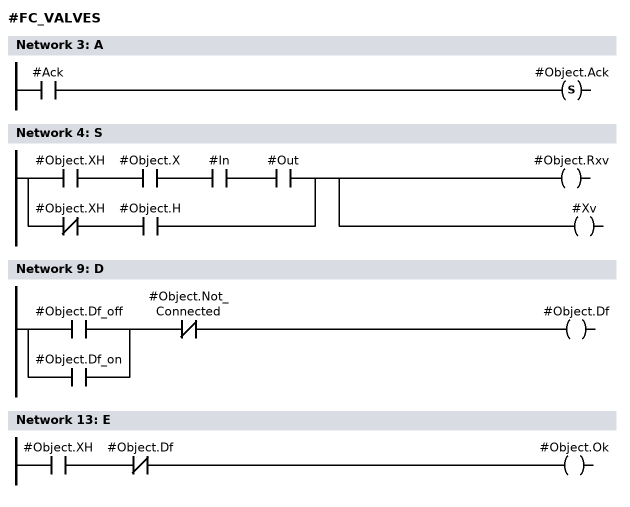
   RUNG wire#powerrail
      Contact( #Ack )
      S_Coil( #Object.Ack )
   END_RUNG
   // the same network as SCL:
   IF #Ack THEN #Object.Ack := TRUE; END_IF;
END_REGION

REGION Network 4: S
   RUNG wire#powerrail
      Contact( #Object.XH )
      Contact( #Object.X )
      Contact( #In )
      Contact( #Out )
      wire#w1
      Coil( #Object.Rxv )
   END_RUNG
   RUNG wire#powerrail
      I_Contact( #Object.XH )
      Contact( #Object.H )
   END_RUNG wire#w1
   RUNG wire#w1
      Coil( #Xv )
   END_RUNG
   // the same network as SCL:
   #Object.Rxv := (#Object.XH AND #Object.X AND #In AND #Out) OR (NOT #Object.XH AND #Object.H);
   #Xv := #Object.Rxv;
END_REGION

REGION Network 5 (STL): M
         A     #Object.XH;
         A     #Object.Rxv;
         S     #Object.H;

         A     #Object.XH;
         AN    #Object.Rxv;
         R     #Object.H;
END_REGION

REGION Network 6 (STL): R
         O(;
         AN    #Object.Inh;
         A     #Zs_on;
         );
         O(;
         A     #Object.Inh;
         A     #Object.Rxv;
         );
         =     #Object.Rzson;


         O(;
         AN    #Object.Inh;
         A     #Zs_off;
         );
         O(;
         A     #Object.Inh;
         AN    #Object.Rxv;
         );
         =     #Object.Rzsoff;


         AN    #In;
         =     #Object.R_in;


         AN    #Out;
         =     #Object.R_out;
END_REGION

REGION Network 7 (STL): D
         A     #Object.Rxv;
         A(;
         A(;
         ON    #Object.Rzson;
         O(;
         A     #Object.Rzsoff;
         A     #Object.Rzson;
         );
         );
         O(;
         A     #Object.Df_on;
         AN    #Object.Ack;
         );
         );
         =     #Temp1;


         CALL  "#FC_TIMER"
         ( Input     := #Temp1,
           Input_RTZ := FALSE,
           Pulse     := "point1secPls",
           RTZ       := FALSE,
           Tbase     := 1,
           Preset1   := #dTime,
           Preset2   := #Object.Gen.Para.Preset_Df_on,
           Time1     := #dTime,
           Time2     := #Object.Internal.Df_on
         );



         AN    #Object.Df_on;
         A(;
         L     #Object.Internal.Df_on;
         L     #Object.Gen.Para.Preset_Df_on;
         ==D;
         );
         JC    FON5;
         JU    FON6;
   FON5: S     #Object.Df_on;


   FON6: A     #Object.Ack;
         JC    FON7;
         JU    FON8;
   FON7: L     0;
         T     #Object.Internal.Df_on;
         R     #Object.Df_on;
   FON8: NOP   0;
END_REGION

REGION Network 8 (STL): d
         AN    #Object.Rxv;
         A(;
         O(;
         ON    #Object.Rzsoff;
         O(;
         A     #Object.Rzsoff;
         A     #Object.Rzson;
         );
         );
         O(;
         A     #Object.Df_off;
         AN    #Object.Ack;
         );
         );
         =     #Temp2;



         CALL  "#FC_TIMER"
         ( Input     := #Temp2,
           Input_RTZ := FALSE,
           Pulse     := "point1secPls",
           RTZ       := FALSE,
           Tbase     := 1,
           Preset1   := #dTime,
           Preset2   := #Object.Gen.Para.Preset_Df_off,
           Time1     := #dTime,
           Time2     := #Object.Internal.Df_off
         );


         AN    #Object.Df_off;
         A(;
         L     #Object.Internal.Df_off;
         L     #Object.Gen.Para.Preset_Df_off;
         ==D;
         );
         JC    FOF5;
         JU    FOF6;
   FOF5: S     #Object.Df_off;


   FOF6: A     #Object.Ack;
         JC    FOF7;
         JU    FOF8;
   FOF7: L     0;
         T     #Object.Internal.Df_off;
         R     #Object.Df_off;
   FOF8: NOP   0;
END_REGION

REGION Network 9: D
   RUNG wire#powerrail
      Contact( #Object.Df_off )
      wire#w1
      I_Contact( #Object.Not_Connected )
      Coil( #Object.Df )
   END_RUNG
   RUNG wire#powerrail
      Contact( #Object.Df_on )
   END_RUNG wire#w1
   // the same network as SCL:
   #Object.Df := (#Object.Df_off OR #Object.Df_on) AND NOT #Object.Not_Connected;
END_REGION

REGION Network 10 (STL): C
         A     #Object.Rxv;
         =     #Object.Internal.X_re_counter;

         CALL  "#FC_COUNTER"
         ( Input    := #Object.Internal.X_re_counter,
           Fr_input := #Object.Internal.Re_counter,
           Raz      := #Object.Raz_Fct_Run,
           Count    := #Object.C_run
         );
END_REGION

REGION Network 11 (STL): T
         CALL  "#FC_TIMER"
         ( Input     := #Object.Internal.X_re_counter,
           Input_RTZ := #Object.Raz_Fct_Run,
           Pulse     := "oneSecPls",
           RTZ       := TRUE,
           Tbase     := 1,
           Preset1   := 2073600000,
           Preset2   := #tTime,
           Time1     := #Object.T_run,
           Time2     := #tTime
         );
END_REGION

REGION Network 12 (STL): I
         CALL  "#FC_INH"
         ( Para_inh   := #Object.Gen.Para.Preset_T_exp_inh,
           Object_inh := #Object.Inh,
           Fe_inh     := #Object.Internal.Fe_inh,
           T_inh      := #Object.Internal.T_exp_inh
         );
END_REGION

REGION Network 13: E
   RUNG wire#powerrail
      Contact( #Object.XH )
      I_Contact( #Object.Df )
      Coil( #Object.Ok )
   END_RUNG
   // the same network as SCL:
   #Object.Ok := #Object.XH AND NOT #Object.Df;
END_REGION

REGION Network 14 (STL): Epics State
   // Copy of Auto/Manual mode
         A     #Object.XH;
         =     #sEpics.sAuto;

   // Copy of Inhibition mode
         A     #Object.Inh;
         =     #sEpics.sSim;

   // Copy of Command
         A     #Object.Rxv;
         =     #sEpics.sCmd;

   // Copy of On sensor
         A     #Object.Rzson;
         =     #sEpics.sOn;

   // Copy of Off sensor
         A     #Object.Rzsoff;
         =     #sEpics.sOff;

   // Copy of On fault
         A     #Object.Df_on;
         =     #sEpics.sOnFlt;

   // Copy of Off fault
         A     #Object.Df_off;
         =     #sEpics.sOffFlt;

   // Copy of Faults
         O     #Object.Df_on;
         O     #Object.Df_off;
         =     #sEpics.sFlt;

   // Copy of Command in Auto
         A     #Object.X;
         =     #sEpics.sCmdAuto;

   // Copy of Type
         A     #sNo;
         =     #sEpics.sNO;
END_REGION

REGION Network 15 (STL): Reset Object Commands
         SET;
         R     #Object.Ack;
         R     #Object.Raz_Fct_Run;
END_REGION
END_FUNCTION

FUNCTION "#FC_CONTROL_HEATER" : Void   // FC313, STL
TITLE = Object : Heater
{ S7_Optimized_Access := 'FALSE' }
VERSION : 0.1
BEGIN

REGION Network 1: Initialise of Equipment
         A     "INIT";
         JCN   INIT;
         S     #Object.XH;
   INIT: NOP   0;
END_REGION

REGION Network 2: Epics Commands
   //Set Auto
         A     #cmdEpics.cmdAuto;
         S     #Object.XH;

   // Set Manu
         A     #cmdEpics.cmdMan;
         R     #Object.XH;

   // Set manual command
         A     #cmdEpics.cmdSet;
         S     #Object.H;

   // Reset manual command
         A     #cmdEpics.cmdRst;
         R     #Object.H;

   // Set High limit
         A     #cmdEpics.cmdHL;
         JCN   Epc0;
         L     #cmdEpics.cHL;
         T     #Object.Tt_Max;
   Epc0: NOP   0;

   // Set Low limit
         A     #cmdEpics.cmdLL;
         JCN   Epc1;
         L     #cmdEpics.cLL;
         T     #Object.Tt_Min;
   Epc1: NOP   0;

   EP01: NOP   0;

   // Reset Epics Commands
         R     #cmdEpics.cmdAuto;
         R     #cmdEpics.cmdMan;
         R     #cmdEpics.cmdSet;
         R     #cmdEpics.cmdRst;
         R     #cmdEpics.cmdHL;
         R     #cmdEpics.cmdLL;
END_REGION

REGION Network 3: Data acquisition
   //Input Temperature
         L     #TtA;
         T     #Object.ValueA;

         L     #TtB;
         T     #Object.ValueB;

         L     #TtC;
         T     #Object.ValueC;

         L     #TtD;
         T     #Object.ValueD;

         L     #TtE;
         T     #Object.ValueE;

         L     #TtF;
         T     #Object.ValueF;


   // Termoswitch
         AN    #TS;
         =     #Object.TS;

   // External Command
         A     #ExtCmd;
         =     #Object.R_ExtCmd;

   //Number of Temperature
         L     #Nb_Tt;
         T     #Object.Nb_Tt;
END_REGION

REGION Network 4: Management Thermoswitch
   //ThermoSwitch
   //Timer On
         A     #Object.TS;
         =     #Rec_Ts_On;

         CALL  "#FC_TIMER"
         ( Input     := #Rec_Ts_On,
           Input_RTZ := FALSE,
           Pulse     := "oneSecPls",
           RTZ       := FALSE,
           Tbase     := 1,
           Preset1   := #Object.P_TS_Ton,
           Preset2   := #T_Time,
           Time1     := #Object.TS_Ton,
           Time2     := #T_Time
         );

         L     #Object.TS_Ton;
         L     #Object.P_TS_Ton;
         >=D;
         S     #Object.TS_Calc;

   //Timer Off
         AN    #Object.TS;
         =     #Rec_Ts_Off;

         CALL  "#FC_TIMER"
         ( Input     := #Rec_Ts_Off,
           Input_RTZ := FALSE,
           Pulse     := "oneSecPls",
           RTZ       := FALSE,
           Tbase     := 1,
           Preset1   := #Object.P_TS_Toff,
           Preset2   := #T_Time,
           Time1     := #Object.TS_Toff,
           Time2     := #T_Time
         );

         L     #Object.TS_Toff;
         L     #Object.P_TS_Toff;
         >=D;
         R     #Object.TS_Calc;
END_REGION

REGION Network 5: Equipment Pilot Command
   //Test of number of temperature to SET
         A(;
         L     #Nb_Tt;
         L     1;
         ==I;
         );
         JC    T01S;
         A(;
         L     #Nb_Tt;
         L     2;
         ==I;
         );
         JC    T02S;
         A(;
         L     #Nb_Tt;
         L     3;
         ==I;
         );
         JC    T03S;
         A(;
         L     #Nb_Tt;
         L     4;
         ==I;
         );
         JC    T04S;
         A(;
         L     #Nb_Tt;
         L     5;
         ==I;
         );
         JC    T05S;
         A(;
         L     #Nb_Tt;
         L     6;
         ==I;
         );
         JC    T06S;

         JU    NCS;

   //Set Command
   T06S: A(;
         L     #Object.ValueF;
         L     #Object.Tt_Min;
         <R;
         );
         S     #Object.Pilot;

   T05S: A(;
         L     #Object.ValueE;
         L     #Object.Tt_Min;
         <R;
         );
         S     #Object.Pilot;

   T04S: A(;
         L     #Object.ValueD;
         L     #Object.Tt_Min;
         <R;
         );
         S     #Object.Pilot;

   T03S: A(;
         L     #Object.ValueC;
         L     #Object.Tt_Min;
         <R;
         );
         S     #Object.Pilot;

   T02S: A(;
         L     #Object.ValueB;
         L     #Object.Tt_Min;
         <R;
         );
         S     #Object.Pilot;

   T01S: A(;
         L     #Object.ValueA;
         L     #Object.Tt_Min;
         <R;
         );
         S     #Object.Pilot;

   NCS:  NOP   0;


   //Test of number of temperature to RESET
         A(;
         L     #Nb_Tt;
         L     1;
         ==I;
         );
         JC    T01R;
         A(;
         L     #Nb_Tt;
         L     2;
         ==I;
         );
         JC    T02R;
         A(;
         L     #Nb_Tt;
         L     3;
         ==I;
         );
         JC    T03R;
         A(;
         L     #Nb_Tt;
         L     4;
         ==I;
         );
         JC    T04R;
         A(;
         L     #Nb_Tt;
         L     5;
         ==I;
         );
         JC    T05R;
         A(;
         L     #Nb_Tt;
         L     6;
         ==I;
         );
         JC    T06R;


   //Reset Command
   T06R: A(;
         L     #Object.ValueF;
         L     #Object.Tt_Max;
         >=R;
         );
         R     #Object.Pilot;

   T05R: A(;
         L     #Object.ValueE;
         L     #Object.Tt_Max;
         >=R;
         );
         R     #Object.Pilot;

   T04R: A(;
         L     #Object.ValueD;
         L     #Object.Tt_Max;
         >=R;
         );
         R     #Object.Pilot;

   T03R: A(;
         L     #Object.ValueC;
         L     #Object.Tt_Max;
         >=R;
         );
         R     #Object.Pilot;

   T02R: A(;
         L     #Object.ValueB;
         L     #Object.Tt_Max;
         >=R;
         );
         R     #Object.Pilot;

   T01R: A(;
         L     #Object.ValueA;
         L     #Object.Tt_Max;
         >=R;
         );
         R     #Object.Pilot;
END_REGION

REGION Network 6: External Pilot
   // External Forcage command
         A     #Object.R_ExtCmd;
         JCN   ExtF;
         S     #Object.Pilot;
   ExtF: NOP   0;
END_REGION

REGION Network 7: Delay of Command
   //Timer On
         A(;
         A     #Object.XH;
         A     #Object.X;
         O;
         AN    #Object.XH;
         A     #Object.H;
         );
         AN    #Object.TS_Calc;
         A     #Object.Pilot;
         =     #Rec_Pilot_On;

         CALL  "#FC_TIMER"
         ( Input     := #Rec_Pilot_On,
           Input_RTZ := FALSE,
           Pulse     := "oneSecPls",
           RTZ       := FALSE,
           Tbase     := 1,
           Preset1   := #Object.P_Pilot_Ton,
           Preset2   := #T_Time,
           Time1     := #Object.Pilot_Ton,
           Time2     := #T_Time
         );

         A(;
         L     #Object.Pilot_Ton;
         L     #Object.P_Pilot_Ton;
         >=D;
         );
         =     #Object.Pilot_Calc;

   // Output command
         A     #Object.Pilot_Calc;
         =     #EH;
         =     #Object.R_EH;
END_REGION

REGION Network 8: Auto copy command on the hand control
         A     #Object.XH;
         A     #Object.R_EH;
         S     #Object.H;

         A     #Object.XH;
         AN    #Object.R_EH;
         R     #Object.H;
END_REGION

REGION Network 9: Equipement ok
         A     #Object.XH;
         =     #Object.Ok;
END_REGION

REGION Network 10: Temps d'utilisation
         CALL  "#FC_TIMER"
         ( Input     := #Object.R_EH,
           Input_RTZ := #Object.Raz_Fct_Run,
           Pulse     := "oneSecPls",
           RTZ       := TRUE,
           Tbase     := 1,
           Preset1   := 2073600000,
           Preset2   := #T_Time,
           Time1     := #Object.T_run,
           Time2     := #T_Time
         );
END_REGION

REGION Network 11: Epics State
   // Copy of Auto/Manual mode
         A     #Object.XH;
         =     #sEpics.sAuto;

   // Copy of ThermoSwitch
         A     #Object.TS;
         =     #sEpics.sTsw;

   // Copy of Heater On signal
         A     #Object.R_EH;
         =     #sEpics.sHtrOn;

   // Copy of Command in Auto Mode
         A     #Object.X;
         =     #sEpics.sCmdAuto;

   // Copy of Command
         A(;
         A     #Object.XH;
         A     #Object.X;
         O;
         AN    #Object.XH;
         A     #Object.H;
         );
         =     #sEpics.sCmd;

   // Copy of High Limit
         L     #Object.Tt_Max;
         T     #sEpics.sHL;

   // Copy of Low Limit
         L     #Object.Tt_Min;
         T     #sEpics.sLL;
END_REGION

REGION Network 12: Reset action bool
         SET;
         R     #Object.Raz_Fct_Run;
END_REGION
END_FUNCTION

FUNCTION "#FC_COUNTER" : Void   // FC320, LAD
TITLE = Object : Counter
{ S7_Optimized_Access := 'FALSE' }
AUTHOR : ISIITECH
VERSION : 1.0
// ISIITECH - Counter
// 19.01.2010 version 1.0
BEGIN

REGION Network 1 (STL): C
         A     #Input;
         FP    #Fr_input;
         JCN   COU1;
         L     #Count;
         L     DINT#2000000000;
         >=D;
         JC    COU2;
         L     1;
         L     #Count;
         +D;
         T     #Count;
   COU1: A     #Raz;
         JCN   COU2;
         L     0;
         T     #Count;
   COU2: NOP   0;
END_REGION
END_FUNCTION

FUNCTION "#FC_INH" : Void   // FC322, LAD
TITLE = Inhibition management
{ S7_Optimized_Access := 'FALSE' }
AUTHOR : ISIITECH
VERSION : 1.0
// ISIITECH - Inhibition
// 19.01.2010 version 1.0
BEGIN

REGION Network 1 (STL): E
         A     "INH_BIT";
         S     #Object_inh;

         A     "INH_BIT";
         A     #Object_inh;
         FP    #Fe_inh;
         R     #Object_inh;
END_REGION

REGION Network 2 (STL): I
         A     #Object_inh;
         A(;
         L     #T_inh;
         L     DINT#0;
         >D;
         );
         JC    INH1;
         L     #Para_inh;
         T     #T_inh;
         SET;
         R     #Object_inh;
         JU    INH2;
   INH1: A     "point1secPls";
         JCN   INH2;
         L     #T_inh;
         L     DINT#100;
         -D;
         T     #T_inh;
   INH2: NOP   0;
END_REGION
END_FUNCTION

FUNCTION "#FC_TIMER" : Void   // FC323, LAD
TITLE = Object : Timer
{ S7_Optimized_Access := 'FALSE' }
AUTHOR : ISIITECH
VERSION : 0.1
// ISIITECH - Timer
// 19.01.2010 version 1.0
BEGIN

REGION Network 1 (STL): T
         A     #Input;
         JCN   ST1;
         L     #Time1;
         L     #Preset1;
         <D;
         JCN   ST2;
         A     #Pulse;
         JCN   ST2;
         L     #Time1;
         L     #Tbase;
         +D;
         T     #Time1;
         JU    ST2;
   ST1:  NOP   0;
   ST2:  NOP   0;



         A(;
         A     #RTZ;
         A     #Input_RTZ;
         );
         O(;
         AN    #Input;
         AN    #RTZ;
         );
         JCN   ST3;
         L     0;
         T     #Time1;
   ST3:  NOP   0;
END_REGION

REGION Network 2 (STL): T
         A     #Input;
         JCN   ST21;
         L     #Time2;
         L     #Preset2;
         <D;
         JCN   ST22;
         A     "point1secPls";
         JCN   ST22;
         L     #Time2;
         L     DINT#100;
         +D;
         T     #Time2;
         JU    ST22;
   ST21: NOP   0;
   ST22: NOP   0;



         A(;
         A     #RTZ;
         A     #Input_RTZ;
         );
         O(;
         AN    #Input;
         AN    #RTZ;
         );
         JCN   ST23;
         L     0;
         T     #Time2;
   ST23: NOP   0;
END_REGION
END_FUNCTION

FUNCTION "INST_VALVES" : Void   // FC406, LAD
TITLE = Instances of Valves
{ S7_Optimized_Access := 'FALSE' }
VERSION : 0.1
BEGIN

REGION Network 1 (STL): GV72
   // Vacuum Gate valve
         CALL  "#FC_VALVES"
         ( In       := TRUE,
           Out      := TRUE,
           sNo      := FALSE,
           Ack      := "Epics_to_PLC".cmdAckn,
           cmdEpics := "Epics_to_PLC".GV72,
           sEpics   := "PLC_to_Epics".GV72,
           Zs_on    := "GV72_open",
           Zs_off   := "GV72_closed",
           Xv       := "GV72_OpenCmd",
           Object   := "#DATA_VALVES".GV72
         );
END_REGION

REGION Network 2 (STL): GV70
   // Vacuum Gate valve
         CALL  "#FC_VALVES"
         ( In       := TRUE,
           Out      := TRUE,
           sNo      := FALSE,
           Ack      := "Epics_to_PLC".cmdAckn,
           cmdEpics := "Epics_to_PLC".GV70,
           sEpics   := "PLC_to_Epics".GV70,
           Zs_on    := "GV70_open",
           Zs_off   := "GV70_closed",
           Xv       := "GV70_OpenCmd",
           Object   := "#DATA_VALVES".GV70
         );
END_REGION

REGION Network 3: Set the valve into automatic mode at startup (IO HMI : Mode Auto (1) / Manu (0))
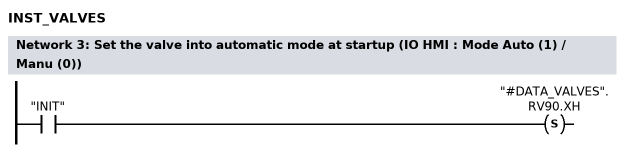
   RUNG wire#powerrail
      Contact( "INIT" )
      S_Coil( "#DATA_VALVES".RV90.XH )
   END_RUNG
   // the same network as SCL:
   IF "INIT" THEN "#DATA_VALVES".RV90.XH := TRUE; END_IF;
END_REGION

REGION Network 4 (STL): RV90
   // Helium release valve
         CALL  "#FC_VALVES"
         ( In       := TRUE,
           Out      := TRUE,
           sNo      := FALSE,
           Ack      := "Epics_to_PLC".cmdAckn,
           cmdEpics := "Epics_to_PLC".RV90,
           sEpics   := "PLC_to_Epics".RV90,
           Zs_on    := "RV90_open",
           Zs_off   := "RV90_closed",
           Xv       := "RV90_OpenCmd",
           Object   := "#DATA_VALVES".RV90
         );
END_REGION
END_FUNCTION

FUNCTION "INST_CONTROL_HEATER" : Void   // FC413, FBD
TITLE = Heater controllers
{ S7_Optimized_Access := 'FALSE' }
AUTHOR : KG
VERSION : 0.1
BEGIN

REGION Network 1 (STL): Init variables
   // Dewar, Electrical Heater
         L     500.0;
         T     #Unused_TT;
         R     #ExtCmd;
END_REGION

REGION Network 2 (STL): EH90 - VB channel 1
   // Dewar, Electrical Heater
         L     2;
         T     "#DATA_HEATERS".EH90.P_TS_Ton;
         T     "#DATA_HEATERS".EH90.P_Pilot_Ton;
         L     5;
         T     "#DATA_HEATERS".EH90.P_TS_Toff;

         SET;
         A     "IOC2PLC".TT900_VALID;
         A     "EPICS_COMM_OK";
         =     #TS;

   // Force the heater ON when the temperature data is not valid
   // (TS = FALSE). The heater will be turned on for 30 s and TS
   // will be forced TRUE for 30 s. This will hopefully raise the
   // temperature enough for Pt100 to be in range (>73 K)
         SET;
         AN    #TS;
         A(;
         A     "#DATA_HEATERS".EH90.XH;
         A     "#DATA_HEATERS".EH90.X;
         O;
         AN    "#DATA_HEATERS".EH90.XH;
         A     "#DATA_HEATERS".EH90.H;
         );
         =     #ExtCmdTrig;
         CALL  TP, "IEC_Timer_EH90_DB"
         ( IN := #ExtCmdTrig,
           PT := T#30s,
           Q  := #ExtCmd,
           ET := #tmp_et
         );
         A     #ExtCmd;
         S     #TS;

         CALL  "#FC_CONTROL_HEATER"
         ( TtA      := "IOC2PLC".TT900,
           TtB      := #Unused_TT,
           TtC      := #Unused_TT,
           TtD      := #Unused_TT,
           TtE      := #Unused_TT,
           TtF      := #Unused_TT,
           Nb_Tt    := 1,
           TS       := #TS,
           ExtCmd   := #ExtCmd,
           cmdEpics := "Epics_to_PLC".EH90,
           EH       := "voie 1 chaufferette BV",
           sEpics   := "PLC_to_Epics".EH90,
           Object   := "#DATA_HEATERS".EH90
         );
END_REGION

REGION Network 3 (STL): EH93-96 - VB channel 2
   // Dewar, Electrical Heater
         L     2;
         T     "#DATA_HEATERS"."EH93-96".P_TS_Ton;
         T     "#DATA_HEATERS"."EH93-96".P_Pilot_Ton;
         L     5;
         T     "#DATA_HEATERS"."EH93-96".P_TS_Toff;

         SET;
         A     "IOC2PLC".TT930_VALID;
         A     "IOC2PLC".TT940_VALID;
         A     "IOC2PLC".TT950_VALID;
         A     "IOC2PLC".TT960_VALID;
         A     "EPICS_COMM_OK";
         =     #TS;

   // Force the heater ON when the temperature data is not valid
   // (TS = FALSE). The heater will be turned on for 30 s and TS
   // will be forced TRUE for 30 s. This will hopefully raise the
   // temperature enough for Pt100 to be in range (>73 K)
         SET;
         AN    #TS;
         A(;
         A     "#DATA_HEATERS"."EH93-96".XH;
         A     "#DATA_HEATERS"."EH93-96".X;
         O;
         AN    "#DATA_HEATERS"."EH93-96".XH;
         A     "#DATA_HEATERS"."EH93-96".H;
         );
         =     #ExtCmdTrig;
         CALL  TP , "IEC_Timer_EH93-96_DB"
         ( IN := #ExtCmdTrig,
           PT := T#30s,
           Q  := #ExtCmd,
           ET := #tmp_et
         );
         A     #ExtCmd;
         S     #TS;

         CALL  "#FC_CONTROL_HEATER"
         ( TtA      := "IOC2PLC".TT930,
           TtB      := "IOC2PLC".TT940,
           TtC      := "IOC2PLC".TT950,
           TtD      := "IOC2PLC".TT960,
           TtE      := #Unused_TT,
           TtF      := #Unused_TT,
           Nb_Tt    := 4,
           TS       := #TS,
           ExtCmd   := #ExtCmd,
           cmdEpics := "Epics_to_PLC"."EH93-96",
           EH       := "voie 2 chaufferette BV",
           sEpics   := "PLC_to_Epics"."EH93-96",
           Object   := "#DATA_HEATERS"."EH93-96"
         );
END_REGION

REGION Network 4 (STL): EH63_64_70 - VB channel 3
   // Dewar, Electrical Heater
         L     2;
         T     "#DATA_HEATERS"."EH63-70".P_TS_Ton;


         T     "#DATA_HEATERS"."EH63-70".P_Pilot_Ton;
         L     5;
         T     "#DATA_HEATERS"."EH63-70".P_TS_Toff;

         SET;
         A     "IOC2PLC".TT630_VALID;
         A     "IOC2PLC".TT640_VALID;
         A     "IOC2PLC".TT700_VALID;
         A     "EPICS_COMM_OK";
         =     #TS;
   // Force the heater ON when the temperature data is not valid
   // (TS = FALSE). The heater will be turned on for 30 s and TS
   // will be forced TRUE for 30 s. This will hopefully raise the
   // temperature enough for Pt100 to be in range (>73 K)
         SET;
         AN    #TS;
         A(;
         A     "#DATA_HEATERS"."EH63-70".XH;
         A     "#DATA_HEATERS"."EH63-70".X;
         O;
         AN    "#DATA_HEATERS"."EH63-70".XH;
         A     "#DATA_HEATERS"."EH63-70".H;
         );
         =     #ExtCmdTrig;
         CALL  TP , "IEC_Timer_EH63-70_DB"
         ( IN := #ExtCmdTrig,
           PT := T#30s,
           Q  := #ExtCmd,
           ET := #tmp_et
         );
         A     #ExtCmd;
         S     #TS;

         CALL  "#FC_CONTROL_HEATER"
         ( TtA      := "IOC2PLC".TT630,
           TtB      := "IOC2PLC".TT640,
           TtC      := "IOC2PLC".TT700,
           TtD      := #Unused_TT,
           TtE      := #Unused_TT,
           TtF      := #Unused_TT,
           Nb_Tt    := 3,
           TS       := #TS,
           ExtCmd   := #ExtCmd,
           cmdEpics := "Epics_to_PLC"."EH63-70",
           EH       := "voie 3 chaufferette BV",
           sEpics   := "PLC_to_Epics"."EH63-70",
           Object   := "#DATA_HEATERS"."EH63-70"
         );
END_REGION

REGION Network 5 (STL): EH61-62 - VB channel 4
   // Dewar, Electrical Heater
         L     2;
         T     "#DATA_HEATERS"."EH61-62".P_TS_Ton;


         T     "#DATA_HEATERS"."EH61-62".P_Pilot_Ton;
         L     5;
         T     "#DATA_HEATERS"."EH61-62".P_TS_Toff;

         SET;
         A     "IOC2PLC".TT610_VALID;
         A     "IOC2PLC".TT620_VALID;
         A     "EPICS_COMM_OK";
         =     #TS;
   // Force the heater ON when the temperature data is not valid
   // (TS = FALSE). The heater will be turned on for 30 s and TS
   // will be forced TRUE for 30 s. This will hopefully raise the
   // temperature enough for Pt100 to be in range (>73 K)
         SET;
         AN    #TS;
         A(;
         A     "#DATA_HEATERS"."EH61-62".XH;
         A     "#DATA_HEATERS"."EH61-62".X;
         O;
         AN    "#DATA_HEATERS"."EH61-62".XH;
         A     "#DATA_HEATERS"."EH61-62".H;
         );
         =     #ExtCmdTrig;
         CALL  TP , "IEC_Timer_EH61-62_DB"
         ( IN := #ExtCmdTrig,
           PT := T#30s,
           Q  := #ExtCmd,
           ET := #tmp_et
         );
         A     #ExtCmd;
         S     #TS;

         CALL  "#FC_CONTROL_HEATER"
         ( TtA      := "IOC2PLC".TT610,
           TtB      := "IOC2PLC".TT620,
           TtC      := #Unused_TT,
           TtD      := #Unused_TT,
           TtE      := #Unused_TT,
           TtF      := #Unused_TT,
           Nb_Tt    := 2,
           TS       := #TS,
           ExtCmd   := #ExtCmd,
           cmdEpics := "Epics_to_PLC"."EH61-62",
           EH       := "voie 4 chaufferette BV",
           sEpics   := "PLC_to_Epics"."EH61-62",
           Object   := "#DATA_HEATERS"."EH61-62"
         );
END_REGION

REGION Network 6 (STL): EH60_67-69 - VB channel 5
   // Dewar, Electrical Heater
         L     2;
         T     "#DATA_HEATERS"."EH60_67-69".P_TS_Ton;


         T     "#DATA_HEATERS"."EH60_67-69".P_Pilot_Ton;
         L     5;
         T     "#DATA_HEATERS"."EH60_67-69".P_TS_Toff;

         SET;
         A     "IOC2PLC".TT600_VALID;
         A     "IOC2PLC".TT670_VALID;
         A     "IOC2PLC".TT680_VALID;
         A     "IOC2PLC".TT690_VALID;
         A     "EPICS_COMM_OK";
         =     #TS;
   // Force the heater ON when the temperature data is not valid
   // (TS = FALSE). The heater will be turned on for 30 s and TS
   // will be forced TRUE for 30 s. This will hopefully raise the
   // temperature enough for Pt100 to be in range (>73 K)
         SET;
         AN    #TS;
         A(;
         A     "#DATA_HEATERS"."EH60_67-69".XH;
         A     "#DATA_HEATERS"."EH60_67-69".X;
         O;
         AN    "#DATA_HEATERS"."EH60_67-69".XH;
         A     "#DATA_HEATERS"."EH60_67-69".H;
         );
         =     #ExtCmdTrig;
         CALL  TP , "IEC_Timer_EH60_67-69_DB"
         ( IN := #ExtCmdTrig,
           PT := T#30s,
           Q  := #ExtCmd,
           ET := #tmp_et
         );
         A     #ExtCmd;
         S     #TS;

         CALL  "#FC_CONTROL_HEATER"
         ( TtA      := "IOC2PLC".TT600,
           TtB      := "IOC2PLC".TT670,
           TtC      := "IOC2PLC".TT680,
           TtD      := "IOC2PLC".TT690,
           TtE      := #Unused_TT,
           TtF      := #Unused_TT,
           Nb_Tt    := 4,
           TS       := #TS,
           ExtCmd   := #ExtCmd,
           cmdEpics := "Epics_to_PLC"."EH60_67-69",
           EH       := "voie 5 chaufferette BV",
           sEpics   := "PLC_to_Epics"."EH60_67-69",
           Object   := "#DATA_HEATERS"."EH60_67-69"
         );
END_REGION

REGION Network 7 (STL): EH97-98 - VB channel 6
   // Dewar, Electrical Heater
         L     2;
         T     "#DATA_HEATERS"."EH97-98".P_TS_Ton;
         T     "#DATA_HEATERS"."EH97-98".P_Pilot_Ton;
         L     5;
         T     "#DATA_HEATERS"."EH97-98".P_TS_Toff;

         SET;
         A     "IOC2PLC".TT970_VALID;
         A     "IOC2PLC".TT980_VALID;
         A     "EPICS_COMM_OK";
         =     #TS;
   // Force the heater ON when the temperature data is not valid
   // (TS = FALSE). The heater will be turned on for 30 s and TS
   // will be forced TRUE for 30 s. This will hopefully raise the
   // temperature enough for Pt100 to be in range (>73 K)
         SET;
         AN    #TS;
         A(;
         A     "#DATA_HEATERS"."EH97-98".XH;
         A     "#DATA_HEATERS"."EH97-98".X;
         O;
         AN    "#DATA_HEATERS"."EH97-98".XH;
         A     "#DATA_HEATERS"."EH97-98".H;
         );
         =     #ExtCmdTrig;
         CALL  TP , "IEC_Timer_EH97-98_DB"
         ( IN := #ExtCmdTrig,
           PT := T#30s,
           Q  := #ExtCmd,
           ET := #tmp_et
         );
         A     #ExtCmd;
         S     #TS;

         CALL  "#FC_CONTROL_HEATER"
         ( TtA      := "IOC2PLC".TT970,
           TtB      := "IOC2PLC".TT980,
           TtC      := #Unused_TT,
           TtD      := #Unused_TT,
           TtE      := #Unused_TT,
           TtF      := #Unused_TT,
           Nb_Tt    := 2,
           TS       := #TS,
           ExtCmd   := #ExtCmd,
           cmdEpics := "Epics_to_PLC"."EH97-98",
           EH       := "voie 6 chaufferette BV",
           sEpics   := "PLC_to_Epics"."EH97-98",
           Object   := "#DATA_HEATERS"."EH97-98"
         );
END_REGION

REGION Network 8 (STL): EH01 - CM channel 1
         L     2;
         T     "#DATA_HEATERS".EH01.P_TS_Ton;
         T     "#DATA_HEATERS".EH01.P_Pilot_Ton;
         L     5;
         T     "#DATA_HEATERS".EH01.P_TS_Toff;

         SET;
         A     "IOC2PLC".TT04_VALID;
         A     "IOC2PLC".TT06_VALID;
         A     "EPICS_COMM_OK";
         =     #TS;

         CALL  "#FC_CONTROL_HEATER"
         ( TtA      := "IOC2PLC".TT04,
           TtB      := "IOC2PLC".TT06,
           TtC      := #Unused_TT,
           TtD      := #Unused_TT,
           TtE      := #Unused_TT,
           TtF      := #Unused_TT,
           Nb_Tt    := 2,
           TS       := #TS,
           ExtCmd   := #ExtCmd,
           cmdEpics := "Epics_to_PLC".EH01,
           EH       := "voie 1 chaufferette CM",
           sEpics   := "PLC_to_Epics".EH01,
           Object   := "#DATA_HEATERS".EH01
         );
END_REGION

REGION Network 9 (STL): EH02 - CM channel 2
         L     2;
         T     "#DATA_HEATERS".EH02.P_TS_Ton;
         T     "#DATA_HEATERS".EH02.P_Pilot_Ton;
         L     5;
         T     "#DATA_HEATERS".EH02.P_TS_Toff;

         SET;
         A     "IOC2PLC".TT05_VALID;
         A     "IOC2PLC".TT07_VALID;
         A     "EPICS_COMM_OK";
         =     #TS;

         CALL  "#FC_CONTROL_HEATER"
         ( TtA      := "IOC2PLC".TT05,
           TtB      := "IOC2PLC".TT07,
           TtC      := #Unused_TT,
           TtD      := #Unused_TT,
           TtE      := #Unused_TT,
           TtF      := #Unused_TT,
           Nb_Tt    := 2,
           TS       := #TS,
           ExtCmd   := #ExtCmd,
           cmdEpics := "Epics_to_PLC".EH02,
           EH       := "voie 2 chaufferette CM",
           sEpics   := "PLC_to_Epics".EH02,
           Object   := "#DATA_HEATERS".EH02
         );
END_REGION

REGION Network 10 (STL): EH10 - CM channel 3
         L     2;
         T     "#DATA_HEATERS".EH10.P_TS_Ton;
         T     "#DATA_HEATERS".EH10.P_Pilot_Ton;
         L     5;
         T     "#DATA_HEATERS".EH10.P_TS_Toff;

         SET;
         A     "IOC2PLC"."CTS:TT10_VALID";
         A     "IOC2PLC"."CTS:TT11_VALID";
         A     "EPICS_COMM_OK";
         =     #TS;

         CALL  "#FC_CONTROL_HEATER"
         ( TtA      := "IOC2PLC"."CTS:TT10",
           TtB      := "IOC2PLC"."CTS:TT11",
           TtC      := #Unused_TT,
           TtD      := #Unused_TT,
           TtE      := #Unused_TT,
           TtF      := #Unused_TT,
           Nb_Tt    := 2,
           TS       := #TS,
           ExtCmd   := #ExtCmd,
           cmdEpics := "Epics_to_PLC".EH10,
           EH       := "voie 3 chaufferette CM",
           sEpics   := "PLC_to_Epics".EH10,
           Object   := "#DATA_HEATERS".EH10
         );
END_REGION

REGION Network 11 (STL): EH20 - CM channel 4
         L     2;
         T     "#DATA_HEATERS".EH20.P_TS_Ton;
         T     "#DATA_HEATERS".EH20.P_Pilot_Ton;
         L     5;
         T     "#DATA_HEATERS".EH20.P_TS_Toff;

         SET;
         A     "IOC2PLC"."CTS:TT20_VALID";
         A     "IOC2PLC"."CTS:TT21_VALID";
         A     "EPICS_COMM_OK";
         =     #TS;

         CALL  "#FC_CONTROL_HEATER"
         ( TtA      := "IOC2PLC"."CTS:TT20",
           TtB      := "IOC2PLC"."CTS:TT21",
           TtC      := #Unused_TT,
           TtD      := #Unused_TT,
           TtE      := #Unused_TT,
           TtF      := #Unused_TT,
           Nb_Tt    := 2,
           TS       := #TS,
           ExtCmd   := #ExtCmd,
           cmdEpics := "Epics_to_PLC".EH20,
           EH       := "voie 4 chaufferette CM",
           sEpics   := "PLC_to_Epics".EH20,
           Object   := "#DATA_HEATERS".EH20
         );
END_REGION

REGION Network 12 (STL): EH918 - CM channel 9
   // Dewar, Electrical Heater
         L     2;
         T     "#DATA_HEATERS"."spare-CM-9".P_TS_Ton;
         T     "#DATA_HEATERS"."spare-CM-9".P_Pilot_Ton;
         L     5;
         T     "#DATA_HEATERS"."spare-CM-9".P_TS_Toff;

         SET;
         A     "IOC2PLC"."CTS:TT20_VALID";
         A     "EPICS_COMM_OK";
         =     #TS;
   // Force the heater ON when the temperature data is not valid
   // (TS = FALSE). The heater will be turned on for 30 s and TS
   // will be forced TRUE for 30 s. This will hopefully raise the
   // temperature enough for Pt100 to be in range (>73 K)
         SET;
         AN    #TS;
         A(;
         A     "#DATA_HEATERS"."spare-CM-9".XH;
         A     "#DATA_HEATERS"."spare-CM-9".X;
         O;
         AN    "#DATA_HEATERS"."spare-CM-9".XH;
         A     "#DATA_HEATERS"."spare-CM-9".H;
         );
         =     #ExtCmdTrig;
         CALL  TP , "IEC_Timer_EH918_DB"
         ( IN := #ExtCmdTrig,
           PT := T#30s,
           Q  := #ExtCmd,
           ET := #tmp_et
         );
         A     #ExtCmd;
         S     #TS;

   _191: CALL  "#FC_CONTROL_HEATER"
         ( TtA      := "IOC2PLC"."CTS:TT20",
           TtB      := #Unused_TT,
           TtC      := #Unused_TT,
           TtD      := #Unused_TT,
           TtE      := #Unused_TT,
           TtF      := #Unused_TT,
           Nb_Tt    := 1,
           TS       := #TS,
           ExtCmd   := #ExtCmd,
           cmdEpics := "Epics_to_PLC"."spare-CM-9",
           EH       := "voie 9 chaufferette CM",
           sEpics   := "PLC_to_Epics"."spare-CM-9",
           Object   := "#DATA_HEATERS"."spare-CM-9"
         );
END_REGION

REGION Network 13 (STL): EH904 - CM channel 11
   // Dewar, Electrical Heater
         L     2;
         T     "#DATA_HEATERS"."spare-CM-11".P_TS_Ton;
         T     "#DATA_HEATERS"."spare-CM-11".P_Pilot_Ton;
         L     5;
         T     "#DATA_HEATERS"."spare-CM-11".P_TS_Toff;

         SET;
         A     "IOC2PLC"."CTS:TT21_VALID";
         A     "EPICS_COMM_OK";
         =     #TS;

   // Force the heater ON when the temperature data is not valid
   // (TS = FALSE). The heater will be turned on for 30 s and TS
   // will be forced TRUE for 30 s. This will hopefully raise the
   // temperature enough for Pt100 to be in range (>73 K)
         SET;
         AN    #TS;
         A(;
         A     "#DATA_HEATERS"."spare-CM-11".XH;
         A     "#DATA_HEATERS"."spare-CM-11".X;
         O;
         AN    "#DATA_HEATERS"."spare-CM-11".XH;
         A     "#DATA_HEATERS"."spare-CM-11".H;
         );
         =     #ExtCmdTrig;
         CALL  TP , "IEC_Timer_EH904_DB"
         ( IN := #ExtCmdTrig,
           PT := T#30s,
           Q  := #ExtCmd,
           ET := #tmp_et
         );
         A     #ExtCmd;
         S     #TS;

         CALL  "#FC_CONTROL_HEATER"
         ( TtA      := "IOC2PLC"."CTS:TT21",
           TtB      := #Unused_TT,
           TtC      := #Unused_TT,
           TtD      := #Unused_TT,
           TtE      := #Unused_TT,
           TtF      := #Unused_TT,
           Nb_Tt    := 1,
           TS       := #TS,
           ExtCmd   := #ExtCmd,
           cmdEpics := "Epics_to_PLC"."spare-CM-11",
           EH       := "voie 11 chaufferette CM",
           sEpics   := "PLC_to_Epics"."spare-CM-11",
           Object   := "#DATA_HEATERS"."spare-CM-11"
         );
END_REGION

REGION Network 14 (STL): EH12 - Coupler 1 flange
   // Dewar, Electrical Heater
         L     2;
         T     "#DATA_HEATERS".EH12.P_TS_Ton;
         T     "#DATA_HEATERS".EH12.P_Pilot_Ton;
         L     5;
         T     "#DATA_HEATERS".EH12.P_TS_Toff;

         L     "PLC_to_Epics".TT120.Visu;
         L     0;
         ==I;
         =     #Enable;
         CALL  "#FC_CONTROL_HEATER"
         ( TtA      := "PLC_to_Epics".TT120.Level,
           TtB      := #Unused_TT,
           TtC      := #Unused_TT,
           TtD      := #Unused_TT,
           TtE      := #Unused_TT,
           TtF      := #Unused_TT,
           Nb_Tt    := 1,
           TS       := #Enable,
           ExtCmd   := #ExtCmd,
           cmdEpics := "Epics_to_PLC".EH12,
           EH       := "EH12 Cpl1",
           sEpics   := "PLC_to_Epics".EH12,
           Object   := "#DATA_HEATERS".EH12
         );
END_REGION

REGION Network 15 (STL): EH22 - Coupler 2 flange
   // Dewar, Electrical Heater
         L     2;
         T     "#DATA_HEATERS".EH22.P_TS_Ton;
         T     "#DATA_HEATERS".EH22.P_Pilot_Ton;
         L     5;
         T     "#DATA_HEATERS".EH22.P_TS_Toff;

         L     "PLC_to_Epics".TT220.Visu;
         L     0;
         ==I;
         =     #Enable;
         CALL  "#FC_CONTROL_HEATER"
         ( TtA      := "PLC_to_Epics".TT220.Level,
           TtB      := #Unused_TT,
           TtC      := #Unused_TT,
           TtD      := #Unused_TT,
           TtE      := #Unused_TT,
           TtF      := #Unused_TT,
           Nb_Tt    := 1,
           TS       := #Enable,
           ExtCmd   := #ExtCmd,
           cmdEpics := "Epics_to_PLC".EH22,
           EH       := "EH22 Cpl2",
           sEpics   := "PLC_to_Epics".EH22,
           Object   := "#DATA_HEATERS".EH22
         );
END_REGION
END_FUNCTION

FUNCTION "Manage_HEATERS" : Void   // FC513, LAD
TITLE = Manage the heaters
{ S7_Optimized_Access := 'FALSE' }
AUTHOR : KG
VERSION : 0.1
BEGIN

REGION Network 1: EH12 & EH22 - Coupler flange cavity 1 and 2
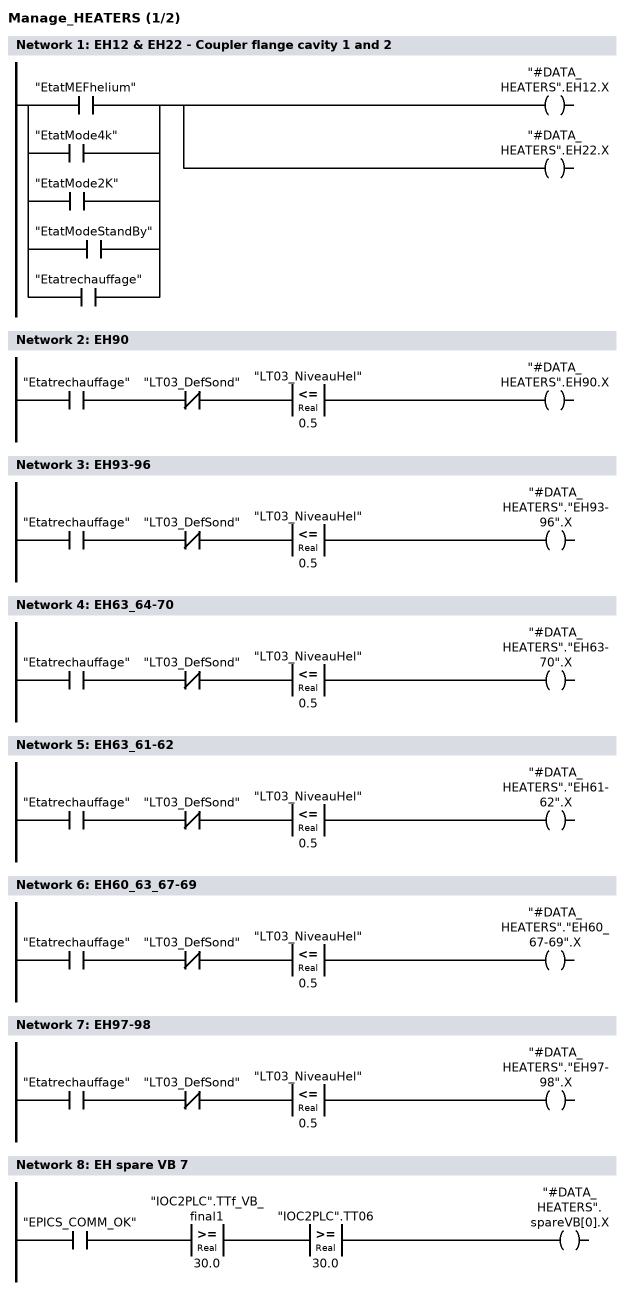
   RUNG wire#powerrail
      Contact( "EtatMEFhelium" )
      wire#w1
      Coil( "#DATA_HEATERS".EH12.X )
   END_RUNG
   RUNG wire#powerrail
      Contact( "EtatMode4k" )
   END_RUNG wire#w1
   RUNG wire#powerrail
      Contact( "EtatMode2K" )
   END_RUNG wire#w1
   RUNG wire#powerrail
      Contact( "EtatModeStandBy" )
   END_RUNG wire#w1
   RUNG wire#powerrail
      Contact( "Etatrechauffage" )
   END_RUNG wire#w1
   RUNG wire#w1
      Coil( "#DATA_HEATERS".EH22.X )
   END_RUNG
   // the same network as SCL:
   "#DATA_HEATERS".EH12.X := "EtatMEFhelium" OR "EtatMode4k" OR "EtatMode2K" OR "EtatModeStandBy" OR "Etatrechauffage";
   "#DATA_HEATERS".EH22.X := "#DATA_HEATERS".EH12.X;
END_REGION

REGION Network 2: EH90
   RUNG wire#powerrail
      Contact( "Etatrechauffage" )
      I_Contact( "LT03_DefSond" )
      { S7_Templates := "SrcType := Real" } LE_Contact(in1 := "LT03_NiveauHel", in2 := 0.5)
      Coil( "#DATA_HEATERS".EH90.X )
   END_RUNG
   // the same network as SCL:
   "#DATA_HEATERS".EH90.X := "Etatrechauffage" AND NOT "LT03_DefSond" AND ("LT03_NiveauHel" <= 0.5);
END_REGION

REGION Network 3: EH93-96
   RUNG wire#powerrail
      Contact( "Etatrechauffage" )
      I_Contact( "LT03_DefSond" )
      { S7_Templates := "SrcType := Real" } LE_Contact(in1 := "LT03_NiveauHel", in2 := 0.5)
      Coil( "#DATA_HEATERS"."EH93-96".X )
   END_RUNG
   // the same network as SCL:
   "#DATA_HEATERS"."EH93-96".X := "Etatrechauffage" AND NOT "LT03_DefSond" AND ("LT03_NiveauHel" <= 0.5);
END_REGION

REGION Network 4: EH63_64-70
   RUNG wire#powerrail
      Contact( "Etatrechauffage" )
      I_Contact( "LT03_DefSond" )
      { S7_Templates := "SrcType := Real" } LE_Contact(in1 := "LT03_NiveauHel", in2 := 0.5)
      Coil( "#DATA_HEATERS"."EH63-70".X )
   END_RUNG
   // the same network as SCL:
   "#DATA_HEATERS"."EH63-70".X := "Etatrechauffage" AND NOT "LT03_DefSond" AND ("LT03_NiveauHel" <= 0.5);
END_REGION

REGION Network 5: EH63_61-62
   RUNG wire#powerrail
      Contact( "Etatrechauffage" )
      I_Contact( "LT03_DefSond" )
      { S7_Templates := "SrcType := Real" } LE_Contact(in1 := "LT03_NiveauHel", in2 := 0.5)
      Coil( "#DATA_HEATERS"."EH61-62".X )
   END_RUNG
   // the same network as SCL:
   "#DATA_HEATERS"."EH61-62".X := "Etatrechauffage" AND NOT "LT03_DefSond" AND ("LT03_NiveauHel" <= 0.5);
END_REGION

REGION Network 6: EH60_63_67-69
   RUNG wire#powerrail
      Contact( "Etatrechauffage" )
      I_Contact( "LT03_DefSond" )
      { S7_Templates := "SrcType := Real" } LE_Contact(in1 := "LT03_NiveauHel", in2 := 0.5)
      Coil( "#DATA_HEATERS"."EH60_67-69".X )
   END_RUNG
   // the same network as SCL:
   "#DATA_HEATERS"."EH60_67-69".X := "Etatrechauffage" AND NOT "LT03_DefSond" AND ("LT03_NiveauHel" <= 0.5);
END_REGION

REGION Network 7: EH97-98
   RUNG wire#powerrail
      Contact( "Etatrechauffage" )
      I_Contact( "LT03_DefSond" )
      { S7_Templates := "SrcType := Real" } LE_Contact(in1 := "LT03_NiveauHel", in2 := 0.5)
      Coil( "#DATA_HEATERS"."EH97-98".X )
   END_RUNG
   // the same network as SCL:
   "#DATA_HEATERS"."EH97-98".X := "Etatrechauffage" AND NOT "LT03_DefSond" AND ("LT03_NiveauHel" <= 0.5);
END_REGION

REGION Network 8: EH spare VB 7
   RUNG wire#powerrail
      Contact( "EPICS_COMM_OK" )
      { S7_Templates := "SrcType := Real" } GE_Contact(in1 := "IOC2PLC".TTf_VB_final1, in2 := 30.0)
      { S7_Templates := "SrcType := Real" } GE_Contact(in1 := "IOC2PLC".TT06, in2 := 30.0)
      Coil( "#DATA_HEATERS".spareVB[0].X )
   END_RUNG
   // the same network as SCL:
   "#DATA_HEATERS".spareVB[0].X := "EPICS_COMM_OK" AND ("IOC2PLC".TTf_VB_final1 >= 30.0) AND ("IOC2PLC".TT06 >= 30.0);
END_REGION

REGION Network 9: EH spare CM 11
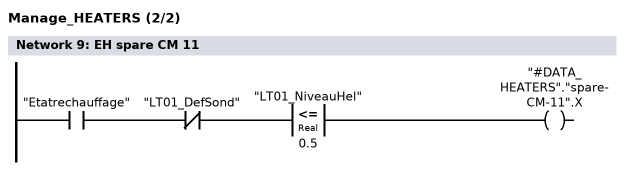
   RUNG wire#powerrail
      Contact( "Etatrechauffage" )
      I_Contact( "LT01_DefSond" )
      { S7_Templates := "SrcType := Real" } LE_Contact(in1 := "LT01_NiveauHel", in2 := 0.5)
      Coil( "#DATA_HEATERS"."spare-CM-11".X )
   END_RUNG
   // the same network as SCL:
   "#DATA_HEATERS"."spare-CM-11".X := "Etatrechauffage" AND NOT "LT01_DefSond" AND ("LT01_NiveauHel" <= 0.5);
END_REGION
END_FUNCTION

FUNCTION "Manage_VALVES" : Void   // FC556, LAD
TITLE = Manage the valves
{ S7_Optimized_Access := 'FALSE' }
AUTHOR : KG
VERSION : 0.1
BEGIN

REGION Network 1: RV90
   // Open the release valve when the pressure is over the threshold
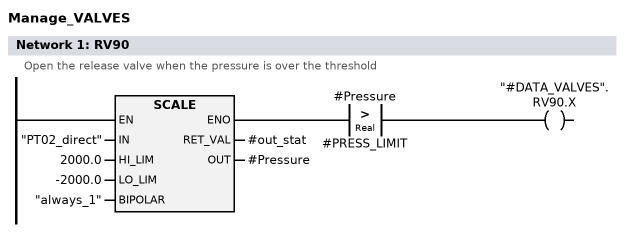
   // ENO of a box is taken as its EN; it also drops when the box reports an error
   #out_stat := SCALE(IN := "PT02_direct",
                      HI_LIM := 2000.0,
                      LO_LIM := -2000.0,
                      BIPOLAR := "always_1",
                      OUT => #Pressure);
   "#DATA_VALVES".RV90.X := #Pressure > #PRESS_LIMIT;
END_REGION
END_FUNCTION

ORGANIZATION_BLOCK "Main"   // OB1, STL
TITLE = "Main Program Sweep (Cycle)"
{ S7_Optimized_Access := 'FALSE' }
VERSION : 0.1
BEGIN

REGION Network 1: Set-up the timing pulse for FC_TIMER
         A     "point1sec";
         AN    "point1secMem";
         =     "point1secPls";
         A     "point1sec";
         =     "point1secMem";

         SET;
         A     "oneSec";
         AN    "oneSecMem";
         =     "oneSecPls";
         A     "oneSec";
         =     "oneSecMem";
END_REGION

REGION Network 2: Get data and commands from Epics IOC
         CALL  "Recv_from_Epics";
         NOP   0;
END_REGION

REGION Network 3
         A     "Graph/manuelle";
         JNB   Label_0;
         CALL  "commande vanne";
   Label_0:NOP   0;
END_REGION

REGION Network 4
         CALL  "NIveau Helium&Pression&vide";
         NOP   0;
END_REGION

REGION Network 5
         CALL  "ACQ_CABTF";
         NOP   0;
END_REGION

REGION Network 6
         AN    "Graph/manuelle";
         JNB   Label_1;
         CALL  "grafcet";
   Label_1:NOP   0;
END_REGION

REGION Network 7
         CALL  "Send_to_Epics";
         NOP   0;
END_REGION

REGION Network 8: Instantiate the heaters control
         CALL  "INST_CONTROL_HEATER";
END_REGION

REGION Network 9: Instantiate the valve control
         CALL  "INST_VALVES";
END_REGION

REGION Network 10: Manage the heaters
         CALL  "Manage_HEATERS";
END_REGION

REGION Network 11: Manage the valves
         CALL  "Manage_VALVES";
END_REGION

REGION Network 12: Clear INIT flag after the first cycle
         SET;
         R     "INIT";
END_REGION

REGION Network 13
         CALL  "UpdateData2HNOSS";
END_REGION

REGION Network 14: Appeler le bloc de diagnostic système / Call system diagnostics block
         CALL  "RSE_FB", "RSE_DB";
END_REGION
END_ORGANIZATION_BLOCK

ORGANIZATION_BLOCK "CYC_INT2"   // OB32, LAD
TITLE = Cyclic_1s / "Cyclic Interrupt"
{ S7_Optimized_Access := 'FALSE' }
AUTHOR : KG
VERSION : 0.1
// Call the PID functionswith 1s interval
   VAR_TEMP   // added for the SCL form of the ladder/FBD networks
      _w1 : Bool;
   END_VAR
BEGIN

REGION Network 1: PID regulator for the LN2 screen cooling (CV60)
